   2290: 'TT426 3S BWT TEMP OUT OF RANGE', class Tank Control Warnings, trigger "2062_Warning_Data_BTCS_WARNING_WORD_11" bit 2
   2291: 'TT426 4P BWT TEMP OUT OF RANGE', class Tank Control Warnings, trigger "2062_Warning_Data_BTCS_WARNING_WORD_11" bit 3
   2292: 'TT426 4S BWT TEMP OUT OF RANGE', class Tank Control Warnings, trigger "2062_Warning_Data_BTCS_WARNING_WORD_11" bit 4
   2293: 'TT426 5P BWT TEMP OUT OF RANGE', class Tank Control Warnings, trigger "2062_Warning_Data_BTCS_WARNING_WORD_11" bit 5
   2294: 'TT426 5S BWT TEMP OUT OF RANGE', class Tank Control Warnings, trigger "2062_Warning_Data_BTCS_WARNING_WORD_11" bit 6
   2295: 'TT426 6P BWT TEMP OUT OF RANGE', class Tank Control Warnings, trigger "2062_Warning_Data_BTCS_WARNING_WORD_11" bit 7
   2296: 'LT422 6S TANK LEVEL HIGH', class Tank Control Warnings, trigger "2062_Warning_Data_BTCS_WARNING_WORD_11" bit 8
   2297: 'LT422 6S TANK LEVEL LOW', class Tank Control Warnings, trigger "2062_Warning_Data_BTCS_WARNING_WORD_11" bit 9
   2298: 'LT422 APT TANK LEVEL HIGH', class Tank Control Warnings, trigger "2062_Warning_Data_BTCS_WARNING_WORD_11" bit 10
   2299: 'LT422 APT TANK LEVEL LOW', class Tank Control Warnings, trigger "2062_Warning_Data_BTCS_WARNING_WORD_11" bit 11
   2300: 'TT426 FPT BWT TEMP OUT OF RANGE', class Tank Control Warnings, trigger "2062_Warning_Data_BTCS_WARNING_WORD_11" bit 12
   2301: 'TT426 1P BWT TEMP OUT OF RANGE', class Tank Control Warnings, trigger "2062_Warning_Data_BTCS_WARNING_WORD_11" bit 13
   2302: 'TT426 1S BWT TEMP OUT OF RANGE', class Tank Control Warnings, trigger "2062_Warning_Data_BTCS_WARNING_WORD_11" bit 14
   2303: 'TT426 2P BWT TEMP OUT OF RANGE', class Tank Control Warnings, trigger "2062_Warning_Data_BTCS_WARNING_WORD_11" bit 15
   2304: 'FIT417 3S USD OUT OF RANGE', class Tank Control Warnings, trigger "2062_Warning_Data_BTCS_WARNING_WORD_12" bit 0
   2305: 'FIT418 4P USD OUT OF RANGE', class Tank Control Warnings, trigger "2062_Warning_Data_BTCS_WARNING_WORD_12" bit 1
   2306: 'FIT417 4S USD OUT OF RANGE', class Tank Control Warnings, trigger "2062_Warning_Data_BTCS_WARNING_WORD_12" bit 2
   2307: 'FIT418 5P USD OUT OF RANGE', class Tank Control Warnings, trigger "2062_Warning_Data_BTCS_WARNING_WORD_12" bit 3
   2308: 'FIT417 5S USD OUT OF RANGE', class Tank Control Warnings, trigger "2062_Warning_Data_BTCS_WARNING_WORD_12" bit 4
   2309: 'FIT418 6P USD OUT OF RANGE', class Tank Control Warnings, trigger "2062_Warning_Data_BTCS_WARNING_WORD_12" bit 5
   2310: 'FIT417 6S USD OUT OF RANGE', class Tank Control Warnings, trigger "2062_Warning_Data_BTCS_WARNING_WORD_12" bit 6
   2311: 'FIT417 APT USD OUT OF RANGE', class Tank Control Warnings, trigger "2062_Warning_Data_BTCS_WARNING_WORD_12" bit 7
   2312: 'TT426 6S BWT TEMP OUT OF RANGE', class Tank Control Warnings, trigger "2062_Warning_Data_BTCS_WARNING_WORD_12" bit 8
   2313: 'TT426 APT BWT TEMP OUT OF RANGE', class Tank Control Warnings, trigger "2062_Warning_Data_BTCS_WARNING_WORD_12" bit 9
   2314: 'FIT418 FPT USD OUT OF RANGE', class Tank Control Warnings, trigger "2062_Warning_Data_BTCS_WARNING_WORD_12" bit 10
   2315: 'FIT418 1P USD OUT OF RANGE', class Tank Control Warnings, trigger "2062_Warning_Data_BTCS_WARNING_WORD_12" bit 11
   2316: 'FIT417 1S USD OUT OF RANGE', class Tank Control Warnings, trigger "2062_Warning_Data_BTCS_WARNING_WORD_12" bit 12
   2317: 'FIT418 2P USD OUT OF RANGE', class Tank Control Warnings, trigger "2062_Warning_Data_BTCS_WARNING_WORD_12" bit 13
   2318: 'FIT417 2S USD OUT OF RANGE', class Tank Control Warnings, trigger "2062_Warning_Data_BTCS_WARNING_WORD_12" bit 14
   2319: 'FIT418 3P USD OUT OF RANGE', class Tank Control Warnings, trigger "2062_Warning_Data_BTCS_WARNING_WORD_12" bit 15
   2320: 'FIT419 4S MBG FLOW OUT OF RANGE', class Tank Control Warnings, trigger "2062_Warning_Data_BTCS_WARNING_WORD_13" bit 0
   2321: 'FIT420 5P MBG FLOW OUT OF RANGE', class Tank Control Warnings, trigger "2062_Warning_Data_BTCS_WARNING_WORD_13" bit 1
   2322: 'FIT419 5S MBG FLOW OUT OF RANGE', class Tank Control Warnings, trigger "2062_Warning_Data_BTCS_WARNING_WORD_13" bit 2
   2323: 'FIT420 6P MBG FLOW OUT OF RANGE', class Tank Control Warnings, trigger "2062_Warning_Data_BTCS_WARNING_WORD_13" bit 3
   2324: 'FIT419 6S MBG FLOW OUT OF RANGE', class Tank Control Warnings, trigger "2062_Warning_Data_BTCS_WARNING_WORD_13" bit 4
   2325: 'FIT420 APT MBG FLOW OUT OF RANGE', class Tank Control Warnings, trigger "2062_Warning_Data_BTCS_WARNING_WORD_13" bit 5
   2326: 'PT415 RIO1 DECK IG PRESSURE OUT OF RANGE', class Tank Control Warnings, trigger "2062_Warning_Data_BTCS_WARNING_WORD_13" bit 6
   2327: 'PT415 RIO2 DECK IG PRESSURE OUT OF RANGE', class Tank Control Warnings, trigger "2062_Warning_Data_BTCS_WARNING_WORD_13" bit 7
   2328: 'FIT420 FPT MBG FLOW OUT OF RANGE', class Tank Control Warnings, trigger "2062_Warning_Data_BTCS_WARNING_WORD_13" bit 8
   2329: 'FIT420 1P MBG FLOW OUT OF RANGE', class Tank Control Warnings, trigger "2062_Warning_Data_BTCS_WARNING_WORD_13" bit 9
   2330: 'FIT419 1S MBG FLOW OUT OF RANGE', class Tank Control Warnings, trigger "2062_Warning_Data_BTCS_WARNING_WORD_13" bit 10
   2331: 'FIT420 2P MBG FLOW OUT OF RANGE', class Tank Control Warnings, trigger "2062_Warning_Data_BTCS_WARNING_WORD_13" bit 11
   2332: 'FIT419 2S MBG FLOW OUT OF RANGE', class Tank Control Warnings, trigger "2062_Warning_Data_BTCS_WARNING_WORD_13" bit 12
   2333: 'FIT420 3P MBG FLOW OUT OF RANGE', class Tank Control Warnings, trigger "2062_Warning_Data_BTCS_WARNING_WORD_13" bit 13
   2334: 'FIT419 3S MBG FLOW OUT OF RANGE', class Tank Control Warnings, trigger "2062_Warning_Data_BTCS_WARNING_WORD_13" bit 14
   2335: 'FIT420 4P MBG FLOW OUT OF RANGE', class Tank Control Warnings, trigger "2062_Warning_Data_BTCS_WARNING_WORD_13" bit 15
   2336: 'PIT424 RIO4 TANK PRESSURE OUT OF RANGE', class Tank Control Warnings, trigger "2062_Warning_Data_BTCS_WARNING_WORD_14" bit 0
   2337: 'PIT424 RIO5 TANK PRESSURE OUT OF RANGE', class Tank Control Warnings, trigger "2062_Warning_Data_BTCS_WARNING_WORD_14" bit 1
   2338: 'PIT424 RIO6 TANK PRESSURE OUT OF RANGE', class Tank Control Warnings, trigger "2062_Warning_Data_BTCS_WARNING_WORD_14" bit 2
   2339: 'PIT424 RIO7 TANK PRESSURE OUT OF RANGE', class Tank Control Warnings, trigger "2062_Warning_Data_BTCS_WARNING_WORD_14" bit 3
   2340: 'LT422 FPT TANK LEVEL OUT OF RANGE', class Tank Control Warnings, trigger "2062_Warning_Data_BTCS_WARNING_WORD_14" bit 4
   2341: 'LT422 1P TANK LEVEL OUT OF RANGE', class Tank Control Warnings, trigger "2062_Warning_Data_BTCS_WARNING_WORD_14" bit 5
   2342: 'LT422 1S TANK LEVEL OUT OF RANGE', class Tank Control Warnings, trigger "2062_Warning_Data_BTCS_WARNING_WORD_14" bit 6
   2343: 'LT422 2P TANK LEVEL OUT OF RANGE', class Tank Control Warnings, trigger "2062_Warning_Data_BTCS_WARNING_WORD_14" bit 7
   2344: 'PT415 RIO3 DECK IG PRESSURE OUT OF RANGE', class Tank Control Warnings, trigger "2062_Warning_Data_BTCS_WARNING_WORD_14" bit 8
   2345: 'PT415 RIO4 DECK IG PRESSURE OUT OF RANGE', class Tank Control Warnings, trigger "2062_Warning_Data_BTCS_WARNING_WORD_14" bit 9
   2346: 'PT415 RIO5 DECK IG PRESSURE OUT OF RANGE', class Tank Control Warnings, trigger "2062_Warning_Data_BTCS_WARNING_WORD_14" bit 10
   2347: 'PT415 RIO6 DECK IG PRESSURE OUT OF RANGE', class Tank Control Warnings, trigger "2062_Warning_Data_BTCS_WARNING_WORD_14" bit 11
   2348: 'PT415 RIO7 DECK IG PRESSURE OUT OF RANGE', class Tank Control Warnings, trigger "2062_Warning_Data_BTCS_WARNING_WORD_14" bit 12
   2349: 'PIT424 RIO1 TANK PRESSURE OUT OF RANGE', class Tank Control Warnings, trigger "2062_Warning_Data_BTCS_WARNING_WORD_14" bit 13
   2350: 'PIT424 RIO2 TANK PRESSURE OUT OF RANGE', class Tank Control Warnings, trigger "2062_Warning_Data_BTCS_WARNING_WORD_14" bit 14
   2351: 'PIT424 RIO3 TANK PRESSURE OUT OF RANGE', class Tank Control Warnings, trigger "2062_Warning_Data_BTCS_WARNING_WORD_14" bit 15
   2352: 'LT422 6S TANK LEVEL OUT OF RANGE', class Tank Control Warnings, trigger "2062_Warning_Data_BTCS_WARNING_WORD_15" bit 0
   2353: 'LT422 APT TANK LEVEL OUT OF RANGE', class Tank Control Warnings, trigger "2062_Warning_Data_BTCS_WARNING_WORD_15" bit 1
   2354: '600-TX-433 APT O2 MONITOR OUT OF RANGE', class Tank Control Warnings, trigger "2062_Warning_Data_BTCS_WARNING_WORD_15" bit 2
   2355: 'PH426 FPT OUT OF RANGE', class Tank Control Warnings, trigger "2062_Warning_Data_BTCS_WARNING_WORD_15" bit 3
   2356: 'PH426 1P OUT OF RANGE', class Tank Control Warnings, trigger "2062_Warning_Data_BTCS_WARNING_WORD_15" bit 4
   2357: 'PH426 1S OUT OF RANGE', class Tank Control Warnings, trigger "2062_Warning_Data_BTCS_WARNING_WORD_15" bit 5
   2358: 'PH426 2P OUT OF RANGE', class Tank Control Warnings, trigger "2062_Warning_Data_BTCS_WARNING_WORD_15" bit 6
   2359: 'PH426 2S OUT OF RANGE', class Tank Control Warnings, trigger "2062_Warning_Data_BTCS_WARNING_WORD_15" bit 7
   2360: 'LT422 2S TANK LEVEL OUT OF RANGE', class Tank Control Warnings, trigger "2062_Warning_Data_BTCS_WARNING_WORD_15" bit 8
   2361: 'LT422 3P TANK LEVEL OUT OF RANGE', class Tank Control Warnings, trigger "2062_Warning_Data_BTCS_WARNING_WORD_15" bit 9
   2362: 'LT422 3S TANK LEVEL OUT OF RANGE', class Tank Control Warnings, trigger "2062_Warning_Data_BTCS_WARNING_WORD_15" bit 10
   2363: 'LT422 4P TANK LEVEL OUT OF RANGE', class Tank Control Warnings, trigger "2062_Warning_Data_BTCS_WARNING_WORD_15" bit 11
   2364: 'LT422 4S TANK LEVEL OUT OF RANGE', class Tank Control Warnings, trigger "2062_Warning_Data_BTCS_WARNING_WORD_15" bit 12
   2365: 'LT422 5P TANK LEVEL OUT OF RANGE', class Tank Control Warnings, trigger "2062_Warning_Data_BTCS_WARNING_WORD_15" bit 13
   2366: 'LT422 5S TANK LEVEL OUT OF RANGE', class Tank Control Warnings, trigger "2062_Warning_Data_BTCS_WARNING_WORD_15" bit 14
   2367: 'LT422 6P TANK LEVEL OUT OF RANGE', class Tank Control Warnings, trigger "2062_Warning_Data_BTCS_WARNING_WORD_15" bit 15
   2368: 'PH425 6S OUT OF RANGE', class Tank Control Warnings, trigger "2062_Warning_Data_BTCS_WARNING_WORD_16" bit 0
   2369: 'PH426 APT OUT OF RANGE', class Tank Control Warnings, trigger "2062_Warning_Data_BTCS_WARNING_WORD_16" bit 1
   2370: 'DO428 FPT OUT OF RANGE', class Tank Control Warnings, trigger "2062_Warning_Data_BTCS_WARNING_WORD_16" bit 2
   2371: 'DO428 1P OUT OF RANGE', class Tank Control Warnings, trigger "2062_Warning_Data_BTCS_WARNING_WORD_16" bit 3
   2372: 'DO427 1S OUT OF RANGE', class Tank Control Warnings, trigger "2062_Warning_Data_BTCS_WARNING_WORD_16" bit 4
   2373: 'DO428 2P OUT OF RANGE', class Tank Control Warnings, trigger "2062_Warning_Data_BTCS_WARNING_WORD_16" bit 5
   2374: 'DO427 2S OUT OF RANGE', class Tank Control Warnings, trigger "2062_Warning_Data_BTCS_WARNING_WORD_16" bit 6
   2375: 'DO428 3P OUT OF RANGE', class Tank Control Warnings, trigger "2062_Warning_Data_BTCS_WARNING_WORD_16" bit 7
   2376: 'PH426 3P OUT OF RANGE', class Tank Control Warnings, trigger "2062_Warning_Data_BTCS_WARNING_WORD_16" bit 8
   2377: 'PH425 3S OUT OF RANGE', class Tank Control Warnings, trigger "2062_Warning_Data_BTCS_WARNING_WORD_16" bit 9
   2378: 'PH426 4P OUT OF RANGE', class Tank Control Warnings, trigger "2062_Warning_Data_BTCS_WARNING_WORD_16" bit 10
   2379: '', class Tank Control Warnings, trigger "2062_Warning_Data_BTCS_WARNING_WORD_16" bit 11
   2380: 'PH425 4S OUT OF RANGE', class Tank Control Warnings, trigger "2062_Warning_Data_BTCS_WARNING_WORD_16" bit 12
   2381: 'PH426 5P OUT OF RANGE', class Tank Control Warnings, trigger "2062_Warning_Data_BTCS_WARNING_WORD_16" bit 13
   2382: 'PH425 5S OUT OF RANGE', class Tank Control Warnings, trigger "2062_Warning_Data_BTCS_WARNING_WORD_16" bit 14
   2383: 'PH426 6P OUT OF RANGE', class Tank Control Warnings, trigger "2062_Warning_Data_BTCS_WARNING_WORD_16" bit 15
   2384: '', class Tank Control Warnings, trigger "2062_Warning_Data_BTCS_WARNING_WORD_17" bit 0
   2385: '', class Tank Control Warnings, trigger "2062_Warning_Data_BTCS_WARNING_WORD_17" bit 1
   2386: '', class Tank Control Warnings, trigger "2062_Warning_Data_BTCS_WARNING_WORD_17" bit 2
   2387: '', class Tank Control Warnings, trigger "2062_Warning_Data_BTCS_WARNING_WORD_17" bit 3
   2388: '', class Tank Control Warnings, trigger "2062_Warning_Data_BTCS_WARNING_WORD_17" bit 4
   2389: '', class Tank Control Warnings, trigger "2062_Warning_Data_BTCS_WARNING_WORD_17" bit 5
   2390: '', class Tank Control Warnings, trigger "2062_Warning_Data_BTCS_WARNING_WORD_17" bit 6
   2391: '', class Tank Control Warnings, trigger "2062_Warning_Data_BTCS_WARNING_WORD_17" bit 7
   2392: 'DO427 3S OUT OF RANGE', class Tank Control Warnings, trigger "2062_Warning_Data_BTCS_WARNING_WORD_17" bit 8
   2393: 'DO428 4P OUT OF RANGE', class Tank Control Warnings, trigger "2062_Warning_Data_BTCS_WARNING_WORD_17" bit 9
   2394: 'DO427 4S OUT OF RANGE', class Tank Control Warnings, trigger "2062_Warning_Data_BTCS_WARNING_WORD_17" bit 10
   2395: 'DO428 5P OUT OF RANGE', class Tank Control Warnings, trigger "2062_Warning_Data_BTCS_WARNING_WORD_17" bit 11
   2396: 'DO427 5S OUT OF RANGE', class Tank Control Warnings, trigger "2062_Warning_Data_BTCS_WARNING_WORD_17" bit 12
   2397: 'DO428 6P OUT OF RANGE', class Tank Control Warnings, trigger "2062_Warning_Data_BTCS_WARNING_WORD_17" bit 13
   2398: 'DO427 6S OUT OF RANGE', class Tank Control Warnings, trigger "2062_Warning_Data_BTCS_WARNING_WORD_17" bit 14
   2399: 'DO428 APT OUT OF RANGE', class Tank Control Warnings, trigger "2062_Warning_Data_BTCS_WARNING_WORD_17" bit 15

text list "P301 Present": 0..1 'P301 Not Pres'; 1 'P301 Present'

text list "CV312 Present": 0..1 'CV312 Not Pres'; 1 'CV312 Present'

text list "CV431 Present": 0..1 'CV431 Not Pres'; 1 'CV431 Present'

text list "CV432 Present": 0..1 'CV432 Not Pres'; 1 'CV432 Present'

text list "STEP LIST IGG": 1 'Step 001 = Confirm Auto Conditions Ok'; 5 'Step 005 = Wait for Start IGG Command'; 10 'Step 010 = Start E131 (IA Compressor)'; 20 'Step 020 = IA Pressure Within Range (PIT112)'; 30 'Step 030 = CSW Outlet Valves In Position'; 40 'Step 040 = CSW Inlet Valves In Position'; 50 'Step 050 = Start P301 (CSW Pump)'; 60 'Step 060 = CSW Inlet pressure Check'; 70 'Step 070 = Check CV203 Position Closed (N.C.)'; 80 'Step 080 = Start E500 (Fuel Pump)'; 90 'Step 090 = Fuel Pressure Within Range (PIT204)'; 100 'Step 100 = Start E139 (CAB)'; 110 'Step 110 = Start Modulation CV403 (Vent Valve) & Check Setpoint Setting'; 120 'Step 120 = Outlet Pressure Within Range (PIT402)'; 130 'Step 130 = Adjust PIT102 Setpoints'; 140 'Step 140 = Pre BC Start Sequence Delay'; 150 'Step 150 = BC Start Command'; 160 'Step 160 = Wait For Pilot Burner Active Status'; 170 'Step 170 = Adjust Setpoints'; 180 'Step 180 = Wait For Pilot Burner Purge Stage Complete'; 190 'Step 190 = Run Setpoint Ramp For PIT402'; 200 'Step 200 = BC Ramp O2 Command'; 210 'Step 210 = Wait For O2 Level OK'; 220 'Step 220 = Wait For Stop Command'; 300 'Step 300 = Stop Command To BC'; 310 'Step 310 = Wait For Stopping Status From BC'; 320 'Step 320 = Wait For O2 Control Stopped From BC'; 330 'Step 330 = Adjust Setpoints'; 340 'Step 340 = Run Setpoint Ramp Down For PIT402'; 350 'Step 350 = Command Burners Off'; 360 'Step 360 = CV403 To 100% (Fully Open)'; 370 'Step 370 = Adjust Setpoints'; 380 'Step 380 = Stop Combustion Air Blower E139'; 390 'Step 390 = Close CV127 Command To BC'; 400 'Step 400 = Stop Fuel Pump'; 410 'Step 410 = Pre CV203 Close Command Delay'; 420 'Step 420 = Close CV203 Command To BC'; 430 'Step 430 = Stop P301 (CSW Pump)'; 440 'Step 440 = P301 Stopped Delay'; 450 'Step 450 = Cooling Water inlet Valves To Initial Position CV311 = Closed & CV312 = Open'; 460 'Step 460 = CV311 Closed Delay'; 470 'Step 470 = Cooling Water Outlet Valves To Initial Position CV321 = Open & CV322 = Closed'; 480 'Step 480 = CV321 Opened Delay'; 490 'Step 490 = Close CV111 Command To BC'; 500 'Step 500 = Wait For Shutdown Status From BC'

text list "STEP LIST BC": 1 'Step 001 = Confirm Auto Conditions Ok'; 5 'Step 005 = Wait for Start BC Command'; 10 'Step 010 = Open Test Pressure valve CV127'; 20 'Step 020 = Check Pressure PS101'; 30 'Step 030 = CV127 Open Delay #1'; 40 'Step 040 = Check Pressure PS101'; 50 'Step 050 = Close Test Pressure valve CV127'; 60 'Step 060 = Check No Pressure PS101'; 70 'Step 070 = CV127 Closed Delay'; 80 'Step 080 = Check No Pressure PS101'; 90 'Step 090 = Open Test Pressure valve CV127'; 100 'Step 100 = Check Pressure PS101'; 110 'Step 110 = CV127 Open Delay #2'; 120 'Step 120 = Check Pressure PS101'; 130 'Step 130 = Open Pilot Burner Ignition Air Valve CV124'; 140 'Step140 = CV124 Open Delay'; 150 'Step 150 = Check Flow FS123'; 160 'Step 160 = Pilot Flame Ignition Sequence Done OK'; 170 'Step 170 = Wait For IGG Confirmation To Continue'; 180 'Step180 = Open CV114'; 190 'Step 190 = CV114 Open Delay'; 200 'Step 200 = Main Burner Ignition Sequence'; 210 'Step 210 = Check Pressure PIT113'; 220 'Step 220 = Pilot Burner Purge Sequence'; 300 'Step 300 = Confirm Shutting Down'; 310 'Step 310 = CV203 To High O2 Standard Burn Setting'; 320 'Step 320 = CV111 To High O2 Standard Burn Setting'; 330 'Step 330 = Modulation Stopped Confirmation To IGG'; 340 'Step 340 = Wait For Stop Burns Command'; 350 'Step 350 = Close CV206'; 360 'Step 360 = CV206 Close Delay'; 370 'Step 370 = Close CV207'; 380 'Step 380 = CV207 Close Delay'; 390 'Step 390 = Close CV114'; 400 'Step 400 = CV114 Close Delay'; 410 'Step 410 = Close CV215'; 420 'Step 420 = CV215 Close Delay'; 430 'Step 430 = Close CV216'; 440 'Step 440 = CV216 Close Delay'; 450 'Step 450 = Close CV124'; 460 'Step 460 = CV124 Close Delay'; 470 'Step 470 = Check No Flame'; 480 'Step 480 = Burn Stopped Confirmation To IGG'; 490 'Step 490 = Wait For Close CV127 Command'; 500 'Step 500 = Close CV127'; 95 'Step 095 = Confirm CV403 Is Open'; 230 'Step 230 = Wait For Ramp O2 Command'; 240 'Step 240 = Run O2 Ramp'; 250 'Step 250 = Wait For O2 In Specification'; 260 'Step 260 = Write O2 Within Specification Status To IGG'; 270 'Step 270 = Wait For Shutdown Command'; 510 'Step 510 = CV127 Close Delay'; 520 'Step 520 = CV127 Closed Confirmation To IGG'; 525 'Step 525 = Wait For Close CV203 Command'; 530 'Step 530 = Close CV203'; 540 'Step 540 = CV203 Closed Confirmation To IGG'; 550 'Step 550 = Wait For Close CV111 Command'; 560 'Step 560 = Close CV111'; 570 'Step 570 = Shutdown Done Status To IGG'

text list "Mod de functionare motor": 1 'AUTOMATIC PLC'; 0 'LOCAL CABINET'; 2 'MANUAL SCADA'; 3 'MANUAL HMI'; 4 'Necunoscut'

text list "Stari motor": 1 'În pauza de răcire'; 2 'Gata de lucru'; 3 'În functiune'; 4 'În avarie'; 5 'Deconectat'; 6 'Condiţii de start OK'; 7 'Necunoscut'

text list "Mod comanda SP1 Automat": 0 'MANUAL'; 1 'AUTOMATIC'

text list "STATE LIST BTCS": 0 'Initial = Waiting for start'; 1 'Pre-Dwell = Period prior to de-oxygenation'; 2 'De-Ox = De-oxygenation'; 3 'Dwell = Period prior to re-oxygenation'; 4 'Re-Ox = Re-oxygenation'; 5 'Post-Dwell = Settle period'; 6 'Shut Down = System shutting down'

text list "Port Tank": 0 'Deactivated'; 1 'Activated'

text list "STEP LIST BTCS": 0 '00 = Initialising'; 1 '01 = Wait for accept & launch'; 5 '05 = Count to prep gas, 30 Mins from Pre-dwell done'; 10 '10 = Wait for preparing gas confirmation'; 15 '15 = Wait For Pre Dwell Done & Gas Available'; 20 '20 = Close activated tank vent valves'; 25 '25 = Open CV406 Gas to deck valve'; 30 '30 = Open CV407 Block valve 1'; 35 '35 = Open CV411 Block valve 2'; 40 '40 = Close CV409 Blead Valve'; 45 '50 = 15s Time delay'; 50 '50 = Open Activated Tank GTT Valves (Gas To Tank)'; 55 '55 = Wait for O2 @ SP For active tanks for 1 minute'; 60 '60 = Wait For DeOx & DeOx @ SP Times Done'; 70 '70 = Confirm IGG Shutdown'; 75 '75 = Close Activated Tank GTT Valves (Gas To Tank)'; 80 '80 = 30s Time delay'; 85 '85 = Open CV409 Blead Valve'; 90 '90 = Close CV406 Gas to deck valve'; 95 '95 = Close CV407 Block Valve 1'; 100 '100 = Close CV411 Block Valve 2'; 110 '110 = Wait For Dwell Time Done'; 120 '120 = Open All Activated Tank Vent Valves'; 125 '125 = Open CV406 Gas to deck valve'; 130 '130 = Open CV407 Block valve 1'; 135 '135 = Open CV411 Block valve 2'; 140 '140 = Close CV409 Blead Valve'; 145 '150 = 15s Time delay'; 150 '150 = Open Activated Tank GTT Valves (Gas To Tank)'; 155 '155 = Wait for O2 @ SP For active tanks for 1 minute'; 160 '160 = Wait For ReOx & ReOx @ SP Times Done'; 170 '170 = Confirm Gas Deleivery Shutdown'; 175 '175 = Close Activated Tank GTT Valves (Gas To Tank)'; 180 '180 = 30s Time delay'; 185 '185 = Open CV409 Blead Valve'; 190 '190 = Close CV406 Gas to deck valve'; 195 '195 = Close CV407 Block Valve 1'; 200 '200 = Close CV411 Block Valve 2'; 210 '210 = Wait For Dwell Time Done'; 220 '220 = System At Shutdown Goto Initialise'

text list "STEP LIST_GCU": 1 'Step 001 = Confirm Auto Conditions Ok'; 5 'Step 005 = Wait For Tank System State Needing Gas'; 10 'Step 010 = Wait For Prepare Gas Command'; 20 'Step 020 = Run Command To IGG'; 30 'Step 030 = Wait For Running & O2 OK Status From IGG'; 40 'Step 040 = Wait For Supply Gas Command'; 50 'Step 050 = Critical Sensor Check'; 60 'Step 060 = Close CV341'; 70 'Step 070 = CV341 Closed Delay'; 80 'Step 080 = Amend Setpoints'; 90 'Step 090 = Open CV358'; 100 'Step 100 = Start P305 (If Fitted)'; 110 'Step 110 = P305 Started Delay'; 120 'Step 120 = Start P304'; 130 'Step 130 = P304 Started Delay'; 140 'Step 140 = GCU Tank Pre-Fill Delay'; 150 'Step 150 = Fill Sucess Or Fail'; 160 'Step 160 = Stop P304'; 170 'Step 170 = P304 Stopped Delay'; 180 'Step 180 = Stop P305 (If Fitted)'; 190 'Step 190 = P305 Stopped Delay'; 200 'Step 200 = Close CV358'; 210 'Step 210 = CV358 Closed Delay'; 220 'Step 220 = Amend Setpoints'; 230 'Step 230 = Start P303'; 240 'Step 240 = P303 Started Delay'; 250 'Step 250 = Confirm No Alarms'; 260 'Step 260 = Start E400'; 270 'Step 270 = E400 Into Loaded Before Step Time Out (E400 Started Delay)'; 280 'Step 280 = E400 On Load Running Delay'; 290 'Step 290 = CV405 Modulation Start & PIT416 Target Ramp Run'; 300 'Step 300 = Amend Setpoints (Not Currently Required = Re-Check)'; 310 'Step 310 = Wiat For BWTS Status (2=DeOx) or (3=Dwell/ReOx)'; 320 'Step 320 = Open CV401'; 330 'Step 330 = CV401 Opened Delay'; 340 'Step 340 = Pre-Open CV441 Sequence Delay'; 350 'Step 350 = Close CV441'; 360 'Step 360 = CV441 Closed Delay (Done = Jump To Step 410)'; 370 'Step 370 = Close CV401'; 380 'Step 380 = CV401 Closed Delay'; 390 'Step 390 = Open CV441'; 400 'Step 400 = CV441 Opened Delay'; 410 'Step 410 = DeOx/ReOx Valave Configuration Done Sequence Delay'; 420 'Step 420 = Wait For Shutdown Instruction +++RUNNING+++'; 430 'Step 430 = Spare Step (Not Used)'; 440 'Step 440 = Spare Step (Not Used)'; 450 'Step 450 = Open CV405 (Start Of Shutdwon Sequence)'; 460 'Step 460 = CV405 Opened Delay'; 470 'Step 470 = Check CV406 Closed (BWT Control)'; 480 'Step 480 = CV406 Closed Delay'; 490 'Step 490 = Open CV441'; 500 'Step 500 = CV441 Opened Delay'; 510 'Step 510 = Close CV401'; 520 'Step 520 = CV401 Closed Delay'; 530 'Step 530 = Stop E400'; 540 'Step 540 = Stop P303'; 550 'Step 550 = P303 Stopped Delay'; 560 'Step 560 = Wait For PIT416 <0.01bar'; 570 'Step 570 = Open CV341'; 580 'Step 580 = CV341 Opened Delay'; 590 'Step 590 = Tank Drain Time Delay'; 600 'Step 600 = Tank Flush Sequence'; 610 'Step 610 = Post Flush Delay'

text list "P305 Present": 0..1 'P305 Not Pres'; 1 'P305 Present'

text list "GCU_LCL": 0 'TAKE CONTROL'; 1 'RELEASE CONTROL'

text list "ENBL_DSBL": 0 'Disabled'; 1 'Enabled'

text list "GTT_OPS": 0 'Open Active GTT Valves'; 1 'Close Active GTT Valves'

text list "BTCS/BWTC": 0 'Activate'; 1 'Deactivate'

text list "PGC Commissioning": 0 'MEA Tank Changeover'; 1 'Please Wait'

text list "IG Transfer": 0 'Cargo Blanketing Mode'; 1 'Balast Water Treatment Mode'

text list "m³/hr to Nm³/hr": 0 'm³/hr to Nm³/hr Conversion'; 1 'm³/hr Raw Value'

graphic list "IA Compressor": 3 'IA Compressor 01'; 0 'IA Compressor 01'; 1 'IA Compressor 02_1'; 2 'IA Compressor 0_1'

graphic list "New IA Compressor": 0 'Graphic_249'; 1 'Graphic_250'; 2 'Graphic_249'; 3 'Graphic_250'

graphic list "Pump Ani": 1 'Pumpd'; 0 'Pump0'; 1 'Pump1'; 2 'Pump2'; 5 'Pumpd'; 3 'Pump0'; 4 'Pump1'

graphic list "IA Compressor_1": 3 'IA Compressor 01'; 0 'IA Compressor 0_1'; 1 'IA Compressor 02_1'; 2 'IA Compressor 0_1'; 0 'IA Compressor 01'

graphic list "IA Compressor_2": 3 'IA Compressor 01'; 0 'IA Compressor 0_1'; 1 'IA Compressor 02_1'; 2 'IA Compressor 0_1'; 0 'IA Compressor 01'

graphic list "IGGS": 0 'Graphic_3'; 1 'Graphic_140'

graphic list "GCU": 0 'Graphic_150'; 1 'Graphic_150'

graphic list "Process time Banner": 2..5 'Graphic_193'; 1 'Pre Dwell'; 2 'Graphic_193'

graphic list "Water Level Override": 0 'Graphic_217'; 1 'Graphic_218'; 2 'Graphic_217'

graphic list "Tank Process Stage": 0 'Graphic_186'; 1 'Selected'; 2 'De-Oxygenation'; 3 'Graphic_189'; 4 'Graphic_190'; 5 'Graphic_191'; 6 'Graphic_192'; 7 'Graphic_186'; 7 'Tank Manually Disabled'

graphic list "Tank Process Stage_II": 0 'INITIAL STATE'; 1 'Pre Dwell'; 2 'De-Oxygenation'; 3 'Graphic_189'; 4 'Graphic_190'; 5 'Graphic_191'; 6 'Graphic_192'; 7 'Graphic_186'

screen "01 Home" 1280x800, template "Template"
   GraphicView "Graphic view_2" at 118,52 size 317x684; Picture "Graphic_137"
   TextField "HmiScreenItemData_4" at 204,164 size 865x50; Text 'Welcome to Coldharbour Marine'
   TextField "HmiScreenItemData_3" at 194,220 size 896x88; Text 'Ballast Water Treatment System'
   Button "HmiScreenItemData" at 116,50 size 1048x686; TextOn 'Main Index'; TextOff 'Text'
      on Release: function_a2a04561(); ActivateScreen("02 Main Index", 0)
   GraphicView "Graphic view_1" at 444,350 size 449x266; Picture "Graphic_185"
   Button "HmiScreenItemData_16" at 98,47 size 1089x692; TextOn 'Back'; TextOff 'Text'
      on Release: function_a2a04561(); ActivateScreen("Balast Water Treatment Plant", 0)
   Button "Button_1" at 1222,758 size 56x40; TextOff 'Text'; PictureOff "Graphic_286"; Authorization "User administration"
      on Release: StopRuntime(0)

screen "04 Alarm Log" 1280x800, template "Template"
   AlarmView "Alarm view_1" at 8,61 size 1258x665
   Button "HmiScreenItemData_1" at 1,1 size 139x43; TextOn 'Back'; TextOff 'Main Index'
      on Release: ActivateScreen("02 Main Index", 0)
   Button "HmiScreenItemData_2" at 143,1 size 139x43; TextOn 'Back'; TextOff 'Alarm Buffer'
      on Release: ActivateScreen("05 Alarm Buffer", 0)
   Button "HmiScreenItemData_3" at 1124,735 size 139x43; TextOn 'RESET ALARMS'; TextOff 'Reset Alarms'
      on Click: function_d9204949("Alarm view_1")
      on Press: function_b14e0dd5("80_From_HMI_Reset_Alarms", 0)
   Button "HmiScreenItemData_18" at 953,735 size 139x43; TextOn 'Back'; TextOff 'Silence Buzzer'; Authorization "User administration"
      on Press: function_b14e0dd5("80_From_HMI_SLNCE_BZR", 0)
      Appearance <- "80_From_HMI_SLNCE_BZR"
   Button "HmiScreenItemData_4" at 1138,1 size 139x43; TextOn 'I&A Compressor Ok'; TextOff 'Back'
      on Release: function_efd93a16()

screen "03 User Admin" 1280x800, template "Template"
   Button "HmiScreenItemData_1" at 1,1 size 159x51; TextOn 'Back'; TextOff 'Main Index'
      on Release: ActivateScreen("02 Main Index", 0)
   UserView "User view_1" at 0,69 size 1279x730
   Button "HmiScreenItemData_4" at 1153,16 size 126x33; TextOn 'I&A Compressor Ok'; TextOff 'Previous Screen'
      on Release: function_efd93a16()

screen "02 Main Index" 1280x800, template "Template"
   on GenerateScreen: "User_Change"()
   GraphicView "Graphic view_1" at 314,58 size 650x705; Picture "Graphic_115"
   TextField "HmiScreenItemData_16" at 80,95 size 880x30; Text 'BALLAST WATER MANAGEMENT SYSTEM'
   Button "HmiScreenItemData_17" at 320,150 size 160x60; TextOn 'IGG Plant'; TextOff 'IGG Plant'; Authorization "Operate"
      on Release: ActivateScreen("Inert Gas Generator Plant", 0)
   Button "HmiScreenItemData_20" at 800,250 size 160x60; TextOn 'IGG Plant'; TextOff 'Commissioning'; Authorization "Commissioning"
      on Release: ActivateScreen("Commissioning Main Page", 0)
   Button "HmiScreenItemData_1" at 2,2 size 159x51; TextOn 'Back'; TextOff 'Home'
      on Release: ActivateScreen("01 Home", 0)
   Button "HmiScreenItemData_4" at 560,250 size 160x60; TextOn 'IGG Plant'; TextOff 'Air System'; Authorization "Operate"
      on Release: ActivateScreen("Air System", 0)
   Button "HmiScreenItemData_7" at 560,150 size 160x60; TextOn 'IGG Plant'; TextOff 'Fuel System'; Authorization "Operate"
      on Release: ActivateScreen("Fuel System", 0)
   Button "HmiScreenItemData_5" at 80,150 size 160x60; TextOn 'IGG Plant'; TextOff 'IGG Setup'; Authorization "Commissioning"
      on Release: ActivateScreen("Inert Gas Generator Setup", 0)
   Button "Button_1" at 800,650 size 160x60; TextOn 'User Account'; TextOff 'User Administration'; Authorization "User administration"
      on Release: ActivateScreen("03 User Admin", 0)
   Button "HmiScreenItemData_9" at 1147,54 size 125x51; TextOn 'IGG Plant'; TextOff 'Login'
      on Click: function_a2a04561()
      on Release: ActivateScreen("Commissioning Main Page", 0)
   Button "HmiScreenItemData_12" at 1147,2 size 125x51; TextOn 'IGG Plant'; TextOff 'Logout'
      on Release: function_f23ef4c9()
   IOField "I/O field_1" at 991,137 size 266x35; FormatPattern ???????????????????????
      ProcessValue <- "Current User"
   Button "HmiScreenItemData_13" at 560,450 size 160x60; TextOn 'IGG Plant'; TextOff 'Fresh Water System'; Authorization "Operate"
      on Release: ActivateScreen("Fresh Water System", 0)
   Button "HmiScreenItemData_2" at 560,350 size 160x60; TextOn 'IGG Plant'; TextOff 'Cooling System'; Authorization "Operate"
      on Release: ActivateScreen("Cooling System", 0)
   Button "Button_2" at 800,150 size 160x60; TextOn 'User Account'; TextOff 'Alarm Log'; Authorization "Operate"
      on Release: ActivateScreen("04 Alarm Log", 0)
   Button "HmiScreenItemData_6" at 320,250 size 160x60; TextOn 'IGG Plant'; TextOff 'GCU Plant'; Authorization "Operate"
      on Release: ActivateScreen("Inert Gas Conditioning Plant", 0)
   Button "HmiScreenItemData_8" at 80,250 size 160x60; TextOn 'IGG Plant'; TextOff 'GCU Setup'; Authorization "Commissioning"
      on Release: ActivateScreen("Inert Gas Conditioning Setup", 0)
   Button "HmiScreenItemData_10" at 320,350 size 160x60; TextOn 'IGG Plant'; TextOff 'BWT Plant'; Authorization "Operate"
      on Release: ActivateScreen("Balast Water Treatment Plant", 0)
   Button "HmiScreenItemData_11" at 91,575 size 160x60; TextOn 'IGG Plant'; TextOff 'BWT Setup'; Authorization "Operate"
      on Release: ActivateScreen("42 BWT Setup", 0)
      Visibility <- "AlwaysTRUE"
   Button "Button_3" at 560,550 size 160x60; TextOn 'User Account'; TextOff 'IG Transfer Mode'; Authorization "Operate"
      on Release: ActivateScreen("IG Transfer Mode", 0)
   Button "Button_4" at 91,455 size 160x60; TextOn 'User Account'; TextOff 'BTCS Setup & Launch'; Authorization "User administration"
      on Release: ActivateScreen("08 BTCS MAIN", 0)
      Visibility <- "AlwaysTRUE"
   Button "Button_5" at 800,350 size 160x60; TextOn 'User Account'; TextOff 'System Configuration'; Authorization "Commissioning"
      on Release: ActivateScreen("09 Sys Config", 0)
   Button "Button_6" at 80,650 size 400x60; TextOn 'User Account'; TextOff 'BWTS (Balast Water Treatment System) Setup & Launch'; Authorization "User administration"
      on Release: ActivateScreen("07 BWTS MAIN", 0)
      Visibility <- "AlwaysTRUE"
   Button "Button_7" at 560,650 size 160x60; TextOn 'User Account'; TextOff 'PGC System'; Authorization "Operate"
      on Release: ActivateScreen("PGC System", 0)
   Button "Button_8" at 60,411 size 199x29; TextOn 'User Account'; TextOff 'Tank Control System'; Authorization "User administration"
   Button "Button_9" at 80,350 size 160x60; TextOn 'User Account'; TextOff 'BTCS Setup & Launch'; Authorization "Operate"
      on Release: ActivateScreen("Balast Water Treatment Setup", 0)
   Button "Button_10" at 800,450 size 160x60; TextOn 'User Account'; TextOff 'Report Test'; Authorization "User administration"
      on Release: ActivateScreen("Reports", 0)
      Visibility <- "user_group"

screen "IGG Analogue Inputs" 1280x800, template "Template"
   on GenerateScreen: "TitleUpdater"()
   Button "HmiScreenItemData_1" at 1,1 size 150x43; TextOn 'Back'; TextOff 'Commissioning'
      on Release: ActivateScreen("Commissioning Main Page", 0)
   TextField "Text field_82" at 60,150 size 220x22; Text 'PIT-102 - CA Pressure (Pre-Ignition)'
   TextField "Text field_90" at 286,124 size 64x20; Text 'Reading'
   IOField "I/O field_2" at 287,150 size 70x22; FormatPattern 9999; Unit  mBar
      ProcessValue <- "12_AI_Data_PIT102_SCALED(1)"
   TextField "Text field_1" at 359,124 size 68x20; Text 'Low Low'
   IOField "I/O field_1" at 361,150 size 60x22; Authorization "Parameter Change"; FormatPattern 9999
      ProcessValue <- "84_Setpoints_PIT102_Pilot_LowLow"
   TextField "Text field_2" at 442,124 size 37x20; Text 'Low'
   IOField "I/O field_3" at 429,150 size 60x22; Authorization "Parameter Change"; FormatPattern 9999
      ProcessValue <- "84_Setpoints_PIT102_Pilot_Low"
   TextField "Text field_3" at 509,124 size 37x20; Text 'High'
   IOField "I/O field_4" at 497,150 size 60x22; Authorization "Parameter Change"; FormatPattern 9999
      ProcessValue <- "84_Setpoints_PIT102_Pilot_High"
   TextField "Text field_4" at 561,124 size 74x20; Text 'High High'
   IOField "I/O field_5" at 565,150 size 60x22; Authorization "Parameter Change"; FormatPattern 9999
      ProcessValue <- "84_Setpoints_PIT102_Pilot_HighHigh"
   TextField "Text field_5" at 434,100 size 76x20; Text 'Setpoints'
   TextField "Text field_6" at 7,150 size 53x22; Text 'IW112'
   TextField "Text field_7" at 60,270 size 220x22; Text 'TIT-401 - IG Temperature'
   IOField "I/O field_6" at 287,270 size 70x22; FormatPattern s999.9; Unit  °C
      ProcessValue <- "12_AI_Data_TIT401_SCALED"
   IOField "I/O field_7" at 361,270 size 60x22; FormatPattern s999.9
   IOField "I/O field_8" at 429,270 size 60x22; FormatPattern s999.9
   IOField "I/O field_9" at 497,270 size 60x22; Authorization "Parameter Change"; FormatPattern s999.9
      ProcessValue <- "84_Setpoints_TIT401_High"
   IOField "I/O field_10" at 565,270 size 60x22; Authorization "Parameter Change"; FormatPattern s999.9
      ProcessValue <- "84_Setpoints_TIT401_HighHigh"
   TextField "Text field_8" at 7,270 size 53x22; Text 'IW114'
   TextField "Text field_9" at 60,310 size 220x22; Text 'PIT-402 - IG Outlet Pres. (Pre-Ignitn.)'
   IOField "I/O field_11" at 287,310 size 70x22; FormatPattern 9999; Unit  mBar
      ProcessValue <- "12_AI_Data_PIT402_SCALED"
   IOField "I/O field_12" at 361,310 size 60x22; Authorization "Parameter Change"; FormatPattern 9999
      ProcessValue <- "84_Setpoints_PIT402_Pilot_LowLow"
   IOField "I/O field_13" at 429,310 size 60x22; Authorization "Parameter Change"; FormatPattern 9999
      ProcessValue <- "84_Setpoints_PIT402_Pilot_Low"
   IOField "I/O field_14" at 497,310 size 60x22; Authorization "Parameter Change"; FormatPattern 9999
      ProcessValue <- "84_Setpoints_PIT402_Pilot_High"
   IOField "I/O field_15" at 565,310 size 60x22; Authorization "Parameter Change"; FormatPattern 9999
      ProcessValue <- "84_Setpoints_PIT402_Pilot_HighHigh"
   TextField "Text field_10" at 7,310 size 53x22; Text 'IW116'
   TextField "Text field_11" at 60,430 size 220x22; Text 'CV-403 - IG Vent Valve Position Fbk'
   IOField "I/O field_16" at 287,430 size 70x22; FormatPattern 999; Unit  %
      ProcessValue <- "12_AI_Data_CV403_SCALED"
   IOField "I/O field_17" at 361,430 size 60x22; FormatPattern 999
   IOField "I/O field_18" at 429,430 size 60x22; FormatPattern 999
   IOField "I/O field_19" at 497,430 size 60x22; FormatPattern 999
   IOField "I/O field_20" at 565,430 size 60x22; FormatPattern 999
   TextField "Text field_12" at 7,430 size 53x22; Text 'IW118'
   TextField "Text field_13" at 60,470 size 220x22; Text 'CA Blower RPM'
   IOField "I/O field_21" at 287,470 size 70x22; FormatPattern 9999; Unit  RPM
      ProcessValue <- "12_AI_Data_E139_RPM_SCALED"
   IOField "I/O field_22" at 361,470 size 60x22; FormatPattern 9999
   IOField "I/O field_23" at 429,470 size 60x22; FormatPattern 9999
   IOField "I/O field_24" at 497,470 size 60x22; FormatPattern 9999
   IOField "I/O field_25" at 565,470 size 60x22; FormatPattern 9999
   TextField "Text field_14" at 7,470 size 54x22; Text 'IW120'
   TextField "Text field_15" at 61,511 size 220x22; Text 'CA Blower Current'
   IOField "I/O field_26" at 288,511 size 70x22; FormatPattern 999.9; Unit  A
      ProcessValue <- "12_AI_Data_E139_AMPS_SCALED"
   IOField "I/O field_27" at 362,511 size 60x22; FormatPattern 9999
   IOField "I/O field_28" at 430,511 size 60x22; FormatPattern 9999
   TextField "Text field_16" at 8,511 size 54x22; Text 'IW122'
   TextField "Text field_17" at 61,552 size 220x22; Text 'LIT-305 - FW Bulk Tank Level'
   IOField "I/O field_31" at 288,552 size 70x22; FormatPattern s99.9; Unit  %
      ProcessValue <- "12_AI_Data_LIT305_SCALED"
   TextField "Text field_18" at 8,552 size 53x22; Text 'IW124'
   TextField "Text field_19" at 61,592 size 220x22; Text 'Spare'
   IOField "I/O field_36" at 288,592 size 70x22; FormatPattern 9.9; Unit  
      ProcessValue <- "12_AI_Data_R1_SPR_AI_126_SCALED"
   IOField "I/O field_37" at 362,592 size 60x22; FormatPattern 9.9
   IOField "I/O field_38" at 430,592 size 60x22; FormatPattern 9.9
   IOField "I/O field_39" at 498,592 size 60x22; FormatPattern 9.9
   IOField "I/O field_40" at 566,592 size 60x22; FormatPattern 9.9
   TextField "Text field_20" at 8,592 size 53x22; Text 'IW126'
   TextField "Text field_21" at 703,151 size 220x22; Text 'Atmospheric Oxygen 1'
   IOField "I/O field_41" at 930,151 size 70x22; FormatPattern 99.99; Unit %
      ProcessValue <- "12_AI_Data_AT_O2_01_SCALED"
   IOField "I/O field_42" at 1004,151 size 60x22; Authorization "Commissioning"; FormatPattern 99.9
      ProcessValue <- "84_Setpoints_AT_O2_1_LowLow"
   IOField "I/O field_43" at 1072,151 size 60x22; Authorization "Commissioning"; FormatPattern 99.9
      ProcessValue <- "84_Setpoints_AT_O2_1_Low"
   IOField "I/O field_44" at 1140,151 size 60x22; FormatPattern 99.9
   IOField "I/O field_45" at 1208,151 size 60x22; FormatPattern 99.9
   TextField "Text field_22" at 650,151 size 53x22; Text 'IW128'
   TextField "Text field_26" at 928,124 size 64x20; Text 'Reading'
   TextField "Text field_27" at 1001,124 size 68x20; Text 'Low Low'
   TextField "Text field_28" at 1082,124 size 37x20; Text 'Low'
   TextField "Text field_29" at 1150,124 size 37x20; Text 'High'
   TextField "Text field_30" at 1203,124 size 74x20; Text 'High High'
   TextField "Text field_31" at 1076,100 size 76x20; Text 'Setpoints'
   TextField "Text field_57" at 703,192 size 220x22; Text 'TIT-315 - Shell CSW Temperature'
   IOField "I/O field_106" at 930,192 size 70x22; FormatPattern s999.9; Unit  °C
      ProcessValue <- "12_AI_Data_TIT315_SCALED"
   IOField "I/O field_107" at 1004,192 size 60x22; FormatPattern s999.9
   IOField "I/O field_108" at 1072,192 size 60x22; FormatPattern s999.9
   TextField "Text field_58" at 650,192 size 54x22; Text 'IW134'
   TextField "Text field_59" at 703,232 size 220x22; Text 'TIT-319 - Inlet CSW Temperature'
   IOField "I/O field_111" at 930,232 size 70x22; FormatPattern s999.9; Unit  °C
      ProcessValue <- "12_AI_Data_TIT319_SCALED"
   IOField "I/O field_112" at 1004,232 size 60x22; FormatPattern s999.9
   IOField "I/O field_113" at 1072,232 size 60x22; FormatPattern s999.9
   TextField "Text field_60" at 650,232 size 53x22; Text 'IW136'
   TextField "Text field_61" at 703,272 size 220x22; Text 'TIT-360 - Outlet CSW Temperature'
   IOField "I/O field_116" at 930,272 size 70x22; FormatPattern s999.9; Unit  °C
      ProcessValue <- "12_AI_Data_TIT360_SCALED"
   IOField "I/O field_117" at 1004,272 size 60x22; FormatPattern s999.9
   IOField "I/O field_118" at 1072,272 size 60x22; FormatPattern s999.9
   TextField "Text field_62" at 650,272 size 53x22; Text 'IW138'
   TextField "Text field_63" at 703,312 size 220x22; Text 'PIT-359 - Inlet CSW Pressure'
   IOField "I/O field_121" at 930,312 size 70x22; FormatPattern 99.9; Unit  Bar
      ProcessValue <- "12_AI_Data_PIT359_SCALED"
   TextField "Text field_64" at 650,312 size 53x22; Text 'IW140'
   TextField "Text field_41" at 133,124 size 89x20; Text 'Description'
   TextField "Text field_42" at 771,124 size 89x20; Text 'Description'
   TextField "Text field_43" at 17,124 size 37x20; Text 'AI'
   TextField "Text field_44" at 661,124 size 37x20; Text 'AI'
   TextField "Text field_47" at 702,352 size 220x22; Text 'PIT-316 - Outlet CSW Pressure'
   IOField "I/O field_81" at 929,352 size 70x22; FormatPattern 99.9; Unit  Bar
      ProcessValue <- "12_AI_Data_PIT316_SCALED"
   TextField "Text field_48" at 649,352 size 53x22; Text 'IW142'
   IOField "I/O field_109" at 1140,192 size 60x22; Authorization "Parameter Change"; FormatPattern s999.9
      ProcessValue <- "84_Setpoints_TIT315_High"
   IOField "I/O field_110" at 1208,192 size 60x22; Authorization "Parameter Change"; FormatPattern s999.9
      ProcessValue <- "84_Setpoints_TIT315_HighHigh"
   IOField "I/O field_114" at 1140,232 size 60x22; Authorization "Parameter Change"; FormatPattern s999.9
      ProcessValue <- "84_Setpoints_TIT319_High"
   IOField "I/O field_115" at 1208,232 size 60x22; Authorization "Parameter Change"; FormatPattern s999.9
      ProcessValue <- "84_Setpoints_TIT319_HighHigh"
   IOField "I/O field_119" at 1140,272 size 60x22; Authorization "Parameter Change"; FormatPattern s999.9
      ProcessValue <- "84_Setpoints_TIT360_High"
   IOField "I/O field_120" at 1208,272 size 60x22; Authorization "Parameter Change"; FormatPattern s999.9
      ProcessValue <- "84_Setpoints_TIT360_HighHigh"
   IOField "I/O field_124" at 1140,312 size 60x22; Authorization "Parameter Change"; FormatPattern 99.9
      ProcessValue <- "84_Setpoints_PIT359_High"
   IOField "I/O field_125" at 1208,312 size 60x22; Authorization "Parameter Change"; FormatPattern 99.9
      ProcessValue <- "84_Setpoints_PIT359_HighHigh"
   IOField "I/O field_84" at 1139,352 size 60x22; Authorization "Parameter Change"; FormatPattern 99.9
      ProcessValue <- "84_Setpoints_PIT316_High"
   IOField "I/O field_85" at 1207,352 size 60x22; Authorization "Parameter Change"; FormatPattern 99.9
      ProcessValue <- "84_Setpoints_PIT316_HighHigh"
   IOField "I/O field_122" at 1004,312 size 60x22; Authorization "Parameter Change"; FormatPattern 99.9
      ProcessValue <- "84_Setpoints_PIT359_LowLow"
   IOField "I/O field_123" at 1072,312 size 60x22; Authorization "Parameter Change"; FormatPattern 99.9
      ProcessValue <- "84_Setpoints_PIT359_Low"
   IOField "I/O field_82" at 1003,352 size 60x22; Authorization "Parameter Change"; FormatPattern 99.9
      ProcessValue <- "84_Setpoints_PIT316_LowLow"
   IOField "I/O field_83" at 1071,352 size 60x22; Authorization "Parameter Change"; FormatPattern 99.9
      ProcessValue <- "84_Setpoints_PIT316_Low"
   TextField "Text field_52" at 17,91 size 333x26; Text 'IGG Control System PLC (Rack 1)'
   TextField "Text field_54" at 649,719 size 228x62; Text 'Note: CSW = Cooling Sea Water'
   Button "Button_1" at 1160,732 size 100x35; TextOn 'BWTS Digital Inputs.'; TextOff 'Next'
      on Click: ActivateScreen("BC Analogue Inputs", 0)
   TextField "Text field_25" at 60,231 size 220x22; Text 'PIT-102 - CA Pressure (Post-Ignition)'
   IOField "I/O field_52" at 361,231 size 60x22; Authorization "Parameter Change"; FormatPattern 9999
      ProcessValue <- "84_Setpoints_PIT102_Post_LowLow"
   IOField "I/O field_53" at 429,231 size 60x22; Authorization "Parameter Change"; FormatPattern 9999
      ProcessValue <- "84_Setpoints_PIT102_Post_Low"
   IOField "I/O field_54" at 497,231 size 60x22; Authorization "Parameter Change"; FormatPattern 9999
      ProcessValue <- "84_Setpoints_PIT102_Post_High"
   IOField "I/O field_55" at 565,231 size 60x22; Authorization "Parameter Change"; FormatPattern 9999
      ProcessValue <- "84_Setpoints_PIT102_Post_HighHigh"
   TextField "Text field_32" at 7,231 size 53x22; Text 'IW112'
   TextField "Text field_33" at 60,391 size 220x22; Text 'PIT-402 - IG Outlet Pres. (Post-Ignitn)'
   IOField "I/O field_57" at 361,391 size 60x22; Authorization "Parameter Change"; FormatPattern 9999
      ProcessValue <- "84_Setpoints_PIT402_Post_LowLow"
   IOField "I/O field_58" at 429,391 size 60x22; Authorization "Parameter Change"; FormatPattern 9999
      ProcessValue <- "84_Setpoints_PIT402_Post_Low"
   IOField "I/O field_59" at 497,391 size 60x22; Authorization "Parameter Change"; FormatPattern 9999
      ProcessValue <- "84_Setpoints_PIT402_Post_High"
   IOField "I/O field_60" at 565,391 size 60x22; Authorization "Parameter Change"; FormatPattern 9999
      ProcessValue <- "84_Setpoints_PIT402_Post_HighHigh"
   TextField "Text field_34" at 7,391 size 53x22; Text 'IW116'
   TextField "Text field_35" at 61,191 size 220x22; Text 'PIT-102 - CA Pressure (Main)'
   IOField "I/O field_50" at 362,191 size 60x22; Authorization "Parameter Change"; FormatPattern 9999
      ProcessValue <- "84_Setpoints_PIT102_Main_LowLow"
   IOField "I/O field_63" at 430,191 size 60x22; Authorization "Parameter Change"; FormatPattern 9999
      ProcessValue <- "84_Setpoints_PIT102_Main_Low"
   IOField "I/O field_64" at 498,191 size 60x22; Authorization "Parameter Change"; FormatPattern 9999
      ProcessValue <- "84_Setpoints_PIT102_Main_High"
   IOField "I/O field_65" at 566,191 size 60x22; Authorization "Parameter Change"; FormatPattern 9999
      ProcessValue <- "84_Setpoints_PIT102_Main_HighHigh"
   TextField "Text field_36" at 8,191 size 53x22; Text 'IW112'
   TextField "Text field_37" at 61,349 size 220x22; Text 'PIT-402 - IG Outlet Pres. (Main)'
   IOField "I/O field_69" at 362,349 size 60x22; Authorization "Parameter Change"; FormatPattern 9999
      ProcessValue <- "84_Setpoints_PIT402_Main_LowLow"
   IOField "I/O field_70" at 430,349 size 60x22; Authorization "Parameter Change"; FormatPattern 9999
      ProcessValue <- "84_Setpoints_PIT402_Main_Low"
   IOField "I/O field_71" at 498,349 size 60x22; Authorization "Parameter Change"; FormatPattern 9999
      ProcessValue <- "84_Setpoints_PIT402_Main_High"
   IOField "I/O field_72" at 566,349 size 60x22; Authorization "Parameter Change"; FormatPattern 9999
      ProcessValue <- "84_Setpoints_PIT402_Main_HighHigh"
   TextField "Text field_38" at 8,349 size 53x22; Text 'IW116'
   IOField "I/O field_29" at 566,511 size 60x22; FormatPattern 9999
   IOField "I/O field_30" at 499,511 size 60x22; FormatPattern 9999
   IOField "I/O field_32" at 361,552 size 60x22; FormatPattern 9999
   IOField "I/O field_33" at 429,552 size 60x22; FormatPattern 9999
   IOField "I/O field_34" at 565,552 size 60x22; FormatPattern 9999
   IOField "I/O field_35" at 498,552 size 60x22; FormatPattern 9999
   TextField "Text field_39" at 1109,687 size 151x62; Text 'To BC Analogue Inputs'
   AlarmView "Alarm view_1" at 0,777 size 1280x23
   Group "Group" at 455,41 size 373x50
   Button "HmiScreenItemData_8" at 469,45 size 355x40; TextOn 'Back'; TextOff 'Text'
   TextField "Screen title" at 455,41 size 373x50; Text 'Screen title'

